(* Logix 5000 project; controller FV vendor 1 type 14 code 217 rev 31.11; software revision 31.00; part 45 of 63 *)
(* tags used below, declared in another part *)
   CWD : CHECKWORD_FLAGS;
   FV_AV1A : PlantItem;   // AV1A
   FV_AV3 : PlantItem;   // AV3
   FV_AV4A : PlantItem;   // AV4A
   FV_B62 : INT[255];   // RESEED FLG
   FV_B72 : INT[255];   // LNCIP FLG
   FV_B72_O_2_OutputBit : BOOL;
   FV_FV10_TTX01_AI : PlantItem;   // FV10_TTX01
   FV_FV11_TTX01_AI : PlantItem;   // FV11_TTX01
   FV_FV12_TTX01_AI : PlantItem;   // FV12_TTX01
   FV_FV13_TTX01_AI : PlantItem;   // FV13_TTX01
   FV_FV14_TTX01_AI : PlantItem;   // FV14_TTX01
   FV_FV15_TTX01_AI : PlantItem;   // FV15_TTX01
   FV_FV16_TTX01_AI : PlantItem;   // FV16_TTX01
   FV_FV17_TTX01_AI : PlantItem;   // FV17_TTX01
   FV_FV18_TTX01_AI : PlantItem;   // FV18_TTX01
   FV_FV19_TTX01_AI : PlantItem;   // FV19_TTX01
   FV_FV1_TTX01_AI : PlantItem;   // FV1_TTX01
   FV_FV20_TTX01_AI : PlantItem;   // FV20_TTX01
   FV_FV21_TTX01_AI : PlantItem;   // FV21_TTX01
   FV_FV22_TTX01_AI : PlantItem;   // FV22_TTX01
   FV_FV23_TTX01_AI : PlantItem;   // FV23_TTX01
   FV_FV24_TTX01_AI : PlantItem;   // FV24_TTX01
   FV_FV25_TTX01_AI : PlantItem;   // FV25_TTX01
   FV_FV26_TTX01_AI : PlantItem;   // FV26_TTX01
   FV_FV26_TTX02_AI : PlantItem;   // FV26_TTX02
   FV_FV27_TTX01_AI : PlantItem;   // FV27_TTX01
   FV_FV27_TTX02_AI : PlantItem;   // FV27_TTX02
   FV_FV28_TTX01_AI : PlantItem;   // FV28_TTX01
   FV_FV28_TTX02_AI : PlantItem;   // FV28_TTX02
   FV_FV29_TTX01_AI : PlantItem;   // FV29_TTX01
   FV_FV29_TTX02_AI : PlantItem;   // FV29_TTX02
   FV_FV2_TTX01_AI : PlantItem;   // FV2_TTX01
   FV_FV30_TTX01_AI : PlantItem;   // FV30_TTX01
   FV_FV30_TTX02_AI : PlantItem;   // FV30_TTX02
   FV_FV31_TTX01_AI : PlantItem;   // FV31_TTX01
   FV_FV31_TTX02_AI : PlantItem;   // FV31_TTX02
   FV_FV3_TTX01_AI : PlantItem;   // FV3_TTX01
   FV_FV4_TTX01_AI : PlantItem;   // FV4_TTX01
   FV_FV5_TTX01_AI : PlantItem;   // FV5_TTX01
   FV_FV6_TTX01_AI : PlantItem;   // FV6_TTX01
   FV_FV7_TTX01_AI : PlantItem;   // FV7_TTX01
   FV_FV8_TTX01_AI : PlantItem;   // FV8_TTX01
   FV_FV9_TTX01_AI : PlantItem;   // FV9_TTX01
   FV_GLYCOL_AI : PlantItem;   // GLYCOL
   FV_N111 : INT[50];   // FV1, CURRENT FV DATA
   FV_N112 : INT[50];   // FV2, CURRENT FV DATA
   FV_N113 : INT[50];   // FV3, CURRENT FV DATA
   FV_N114 : INT[50];   // FV4, CURRENT FV DATA
   FV_N115 : INT[50];   // FV5, CURRENT FV DATA
   FV_N116 : INT[50];   // FV6, CURRENT FV DATA
   FV_N117 : INT[50];   // FV7, CURRENT FV DATA
   FV_N118 : INT[50];   // FV8, CURRENT FV DATA
   FV_N119 : INT[50];   // FV9, CURRENT FV DATA
   FV_N12 : INT[255];   // SYS_PARMS System Parameter Fil e
   FV_N120 : INT[50];   // FV10, CURRENT FV DATA
   FV_N121 : INT[50];   // FV11, CURRENT FV DATA
   FV_N122 : INT[50];   // FV12, CURRENT FV DATA
   FV_N123 : INT[50];   // FV13, CURRENT FV DATA
   FV_N124 : INT[50];   // FV14, CURRENT FV DATA
   FV_N125 : INT[50];   // FV15, CURRENT FV DATA
   FV_N126 : INT[50];   // FV16, CURRENT FV DATA
   FV_N127 : INT[50];   // FV17, CURRENT FV DATA
   FV_N128 : INT[50];   // FV18, CURRENT FV DATA
   FV_N129 : INT[50];   // FV19, CURRENT FV DATA
   FV_N130 : INT[50];   // FV20, CURRENT FV DATA
   FV_N131 : INT[50];   // FV21, CURRENT FV DATA
   FV_N132 : INT[50];   // FV22, CURRENT FV DATA
   FV_N133 : INT[50];   // FV23, CURRENT FV DATA
   FV_N134 : INT[50];   // FV24, CURRENT FV DATA
   FV_N135 : INT[50];   // FV25, CURRENT FV DATA
   FV_N136 : INT[50];   // YSV1, CURRENT FV DATA
   FV_N137 : INT[50];   // YSV2, CURRENT FV DATA
   FV_N138 : INT[50];   // YSV3, CURRENT FV DATA
   FV_N139 : INT[255];   // YST1
   FV_N140 : INT[255];   // YST2
   FV_N141 : INT[255];   // YSV1 DATA
   FV_N142 : INT[255];   // YSV2 DATA
   FV_N143 : INT[255];   // YSV3 DATA
   FV_N146 : INT[50];   // FV26, CURRENT FV DATA
   FV_N147 : INT[50];   // FV27, CURRENT FV DATA
   FV_N148 : INT[50];   // FV28, CURRENT FV DATA
   FV_N149 : INT[50];   // FV29, CURRENT FV DATA
   FV_N150 : INT[50];   // FV30, CURRENT FV DATA
   FV_N151 : INT[50];   // FV31, CURRENT FV DATA
   FV_N7 : INT[255];   // INTEGER
   FV_N70 : INT[255];   // LNCIP <PC
   FV_N71 : INT[255];   // LNCIP >PC
   FV_PX2 : PlantItem;   // PX2
   FV_PX3 : PlantItem;   // PX3
   FV_SOV1 : PlantItem;   // SOV1
   FV_T73 : TIMER[10];
   FV_TTX_YS_001_AI : PlantItem;   // TTX_YS_001
   FV_TTX_YS_002_AI : PlantItem;   // TTX_YS_002
   FV_YSV1_TTX01_AI : PlantItem;   // YSV1_TTX01
   FV_YSV1_WTX01_AI : PlantItem;   // YSV1_WTX01
   FV_YSV2_TTX01_AI : PlantItem;   // YSV2_TTX01
   FV_YSV2_WTX01_AI : PlantItem;   // YSV2_WTX01
   FV_YSV3_TTX01_AI : PlantItem;   // YSV3_TTX01
   FV_YSV3_WTX01_AI : PlantItem;   // YSV3_WTX01
(* FV_Common, continued *)

ROUTINE FV_LNCIP_CP_36   (* ladder *)
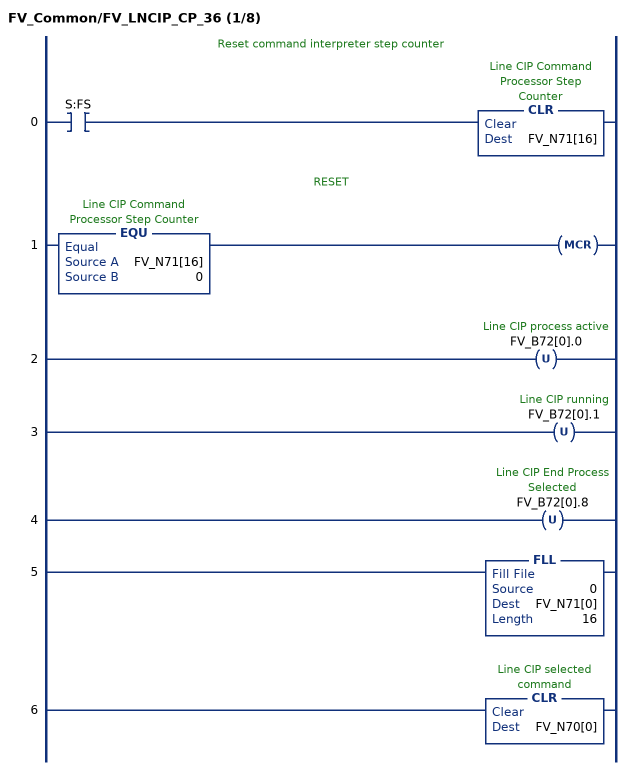
   // Reset command interpreter step counter
   0: XIC(S:FS)CLR(FV_N71[16]);
   // RESET
   1: EQU(FV_N71[16],0)MCR();
   2: OTU(FV_B72[0].0);
   3: OTU(FV_B72[0].1);
   4: OTU(FV_B72[0].8);
   5: FLL(0,FV_N71[0],16);
   6: CLR(FV_N70[0]);
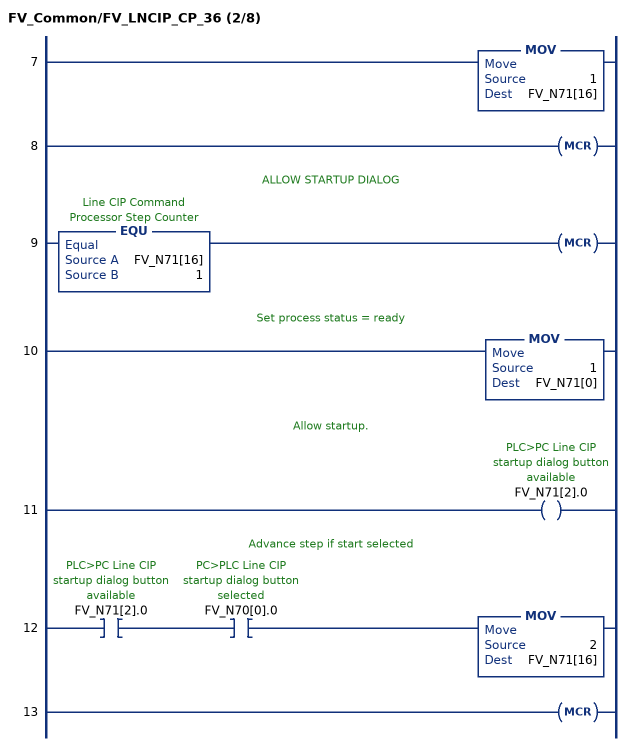
   7: MOV(1,FV_N71[16]);
   8: MCR();
   // ALLOW STARTUP DIALOG
   9: EQU(FV_N71[16],1)MCR();
   // Set process status = ready
   10: MOV(1,FV_N71[0]);
   // Allow startup.
   11: OTE(FV_N71[2].0);
   // Advance step if start selected
   12: XIC(FV_N71[2].0)XIC(FV_N70[0].0)MOV(2,FV_N71[16]);
   13: MCR();
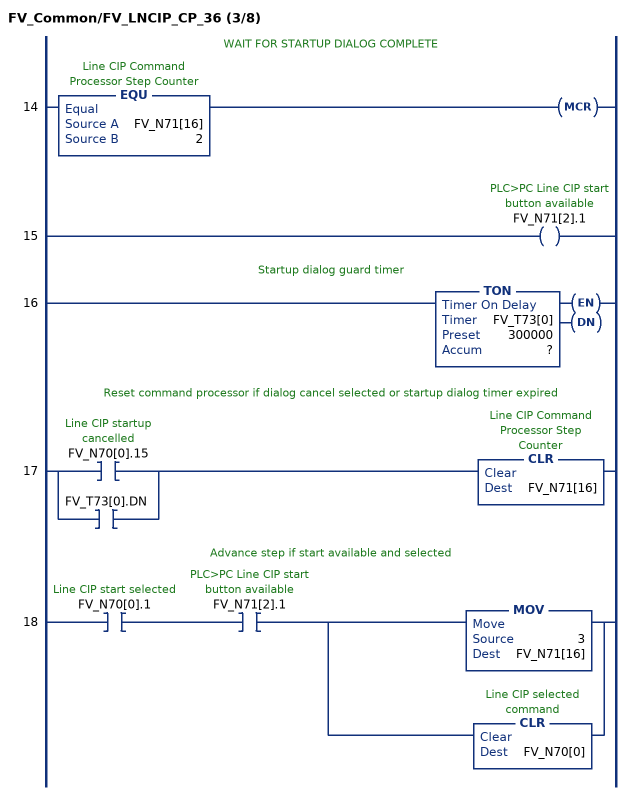
   // WAIT FOR STARTUP DIALOG COMPLETE
   14: EQU(FV_N71[16],2)MCR();
   15: OTE(FV_N71[2].1);
   // Startup dialog guard timer
   16: TON(FV_T73[0],?,?);
   // Reset command processor if dialog cancel selected or startup dialog timer expired
   17: [XIC(FV_N70[0].15) ,XIC(FV_T73[0].DN) ]CLR(FV_N71[16]);
   // Advance step if start available and selected
   18: XIC(FV_N70[0].1)XIC(FV_N71[2].1)[MOV(3,FV_N71[16]) ,CLR(FV_N70[0]) ];
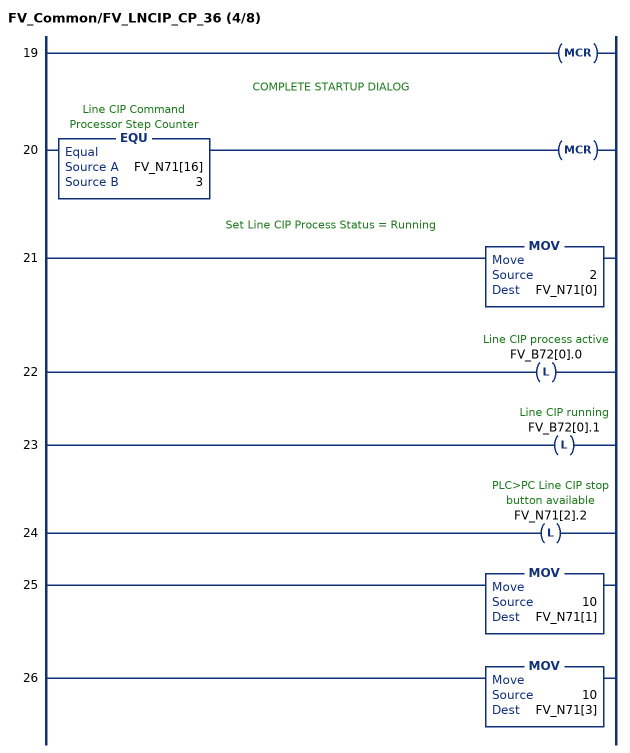
   19: MCR();
   // COMPLETE STARTUP DIALOG
   20: EQU(FV_N71[16],3)MCR();
   // Set Line CIP Process Status = Running
   21: MOV(2,FV_N71[0]);
   22: OTL(FV_B72[0].0);
   23: OTL(FV_B72[0].1);
   24: OTL(FV_N71[2].2);
   25: MOV(10,FV_N71[1]);
   26: MOV(10,FV_N71[3]);
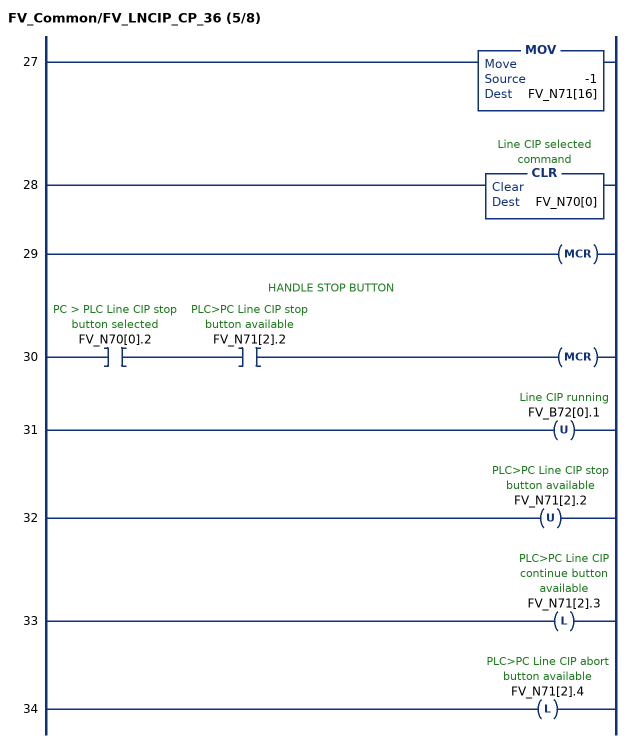
   27: MOV(-1,FV_N71[16]);
   28: CLR(FV_N70[0]);
   29: MCR();
   // HANDLE STOP BUTTON
   30: XIC(FV_N70[0].2)XIC(FV_N71[2].2)MCR();
   31: OTU(FV_B72[0].1);
   32: OTU(FV_N71[2].2);
   33: OTL(FV_N71[2].3);
   34: OTL(FV_N71[2].4);
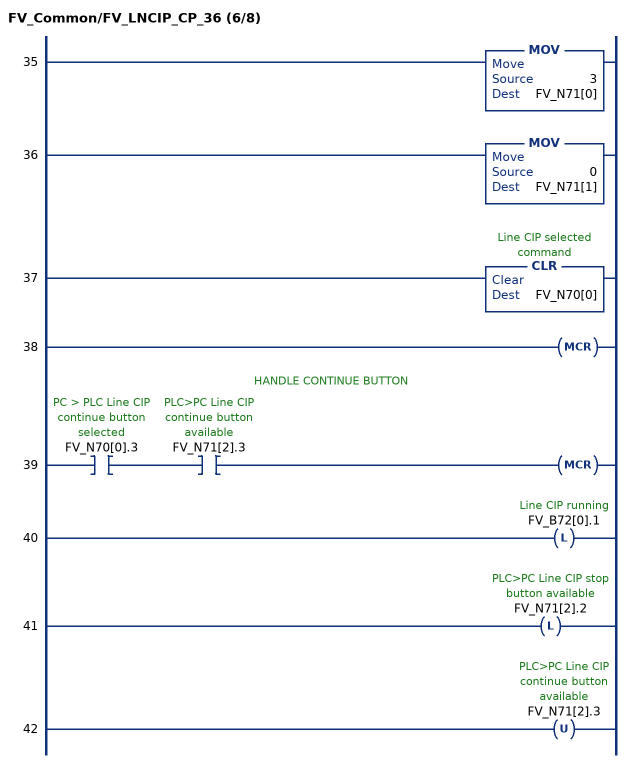
   35: MOV(3,FV_N71[0]);
   36: MOV(0,FV_N71[1]);
   37: CLR(FV_N70[0]);
   38: MCR();
   // HANDLE CONTINUE BUTTON
   39: XIC(FV_N70[0].3)XIC(FV_N71[2].3)MCR();
   40: OTL(FV_B72[0].1);
   41: OTL(FV_N71[2].2);
   42: OTU(FV_N71[2].3);
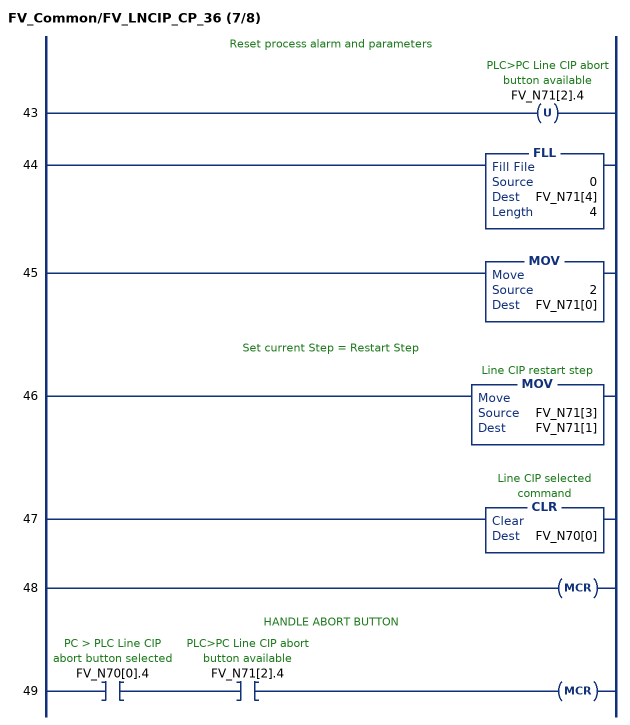
   // Reset process alarm and parameters
   43: OTU(FV_N71[2].4);
   44: FLL(0,FV_N71[4],4);
   45: MOV(2,FV_N71[0]);
   // Set current Step = Restart Step
   46: MOV(FV_N71[3],FV_N71[1]);
   47: CLR(FV_N70[0]);
   48: MCR();
   // HANDLE ABORT BUTTON
   49: XIC(FV_N70[0].4)XIC(FV_N71[2].4)MCR();
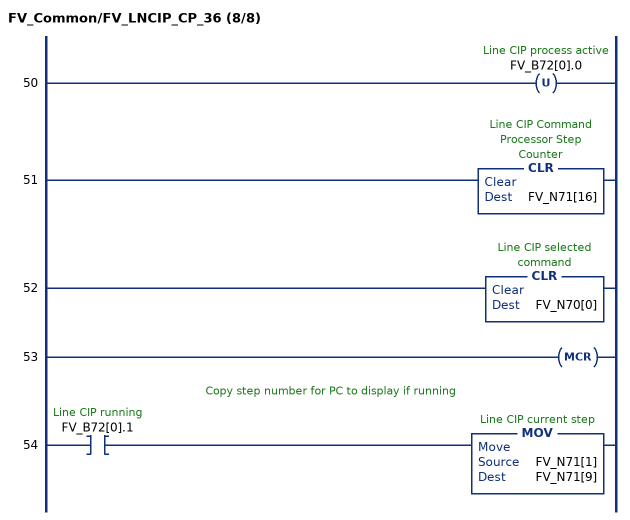
   50: OTU(FV_B72[0].0);
   51: CLR(FV_N71[16]);
   52: CLR(FV_N70[0]);
   53: MCR();
   // Copy step number for PC to display if running
   54: XIC(FV_B72[0].1)MOV(FV_N71[1],FV_N71[9]);
END_ROUTINE

ROUTINE FV_LNCIP_MC_35   (* ladder *)
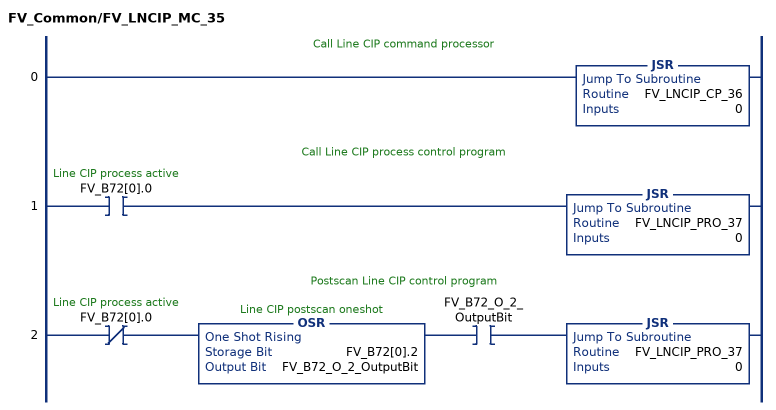
   // Call Line CIP command processor
   0: JSR(FV_LNCIP_CP_36,0);
   // Call Line CIP process control program
   1: XIC(FV_B72[0].0)JSR(FV_LNCIP_PRO_37,0);
   // Postscan Line CIP control program
   2: XIO(FV_B72[0].0)OSR(FV_B72[0].2,FV_B72_O_2_OutputBit)XIC(FV_B72_O_2_OutputBit)JSR(FV_LNCIP_PRO_37,0);
END_ROUTINE

ROUTINE FV_LNCIP_PRO_37   (* ladder *)
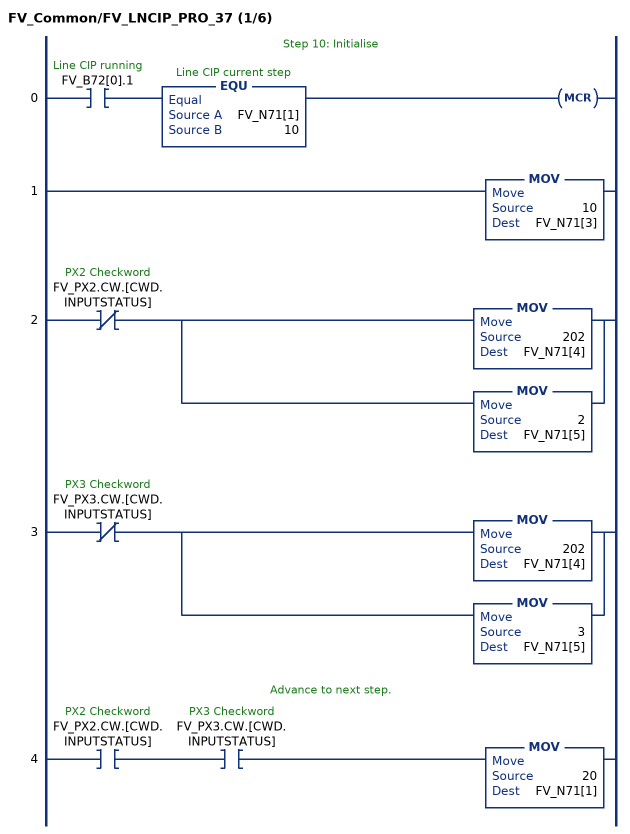
   // Step 10: Initialise
   0: XIC(FV_B72[0].1)EQU(FV_N71[1],10)MCR();
   1: MOV(10,FV_N71[3]);
   2: XIO(FV_PX2.CW.[CWD.INPUTSTATUS])[MOV(202,FV_N71[4]) ,MOV(2,FV_N71[5]) ];
   3: XIO(FV_PX3.CW.[CWD.INPUTSTATUS])[MOV(202,FV_N71[4]) ,MOV(3,FV_N71[5]) ];
   // Advance to next step.
   4: XIC(FV_PX2.CW.[CWD.INPUTSTATUS])XIC(FV_PX3.CW.[CWD.INPUTSTATUS])MOV(20,FV_N71[1]);
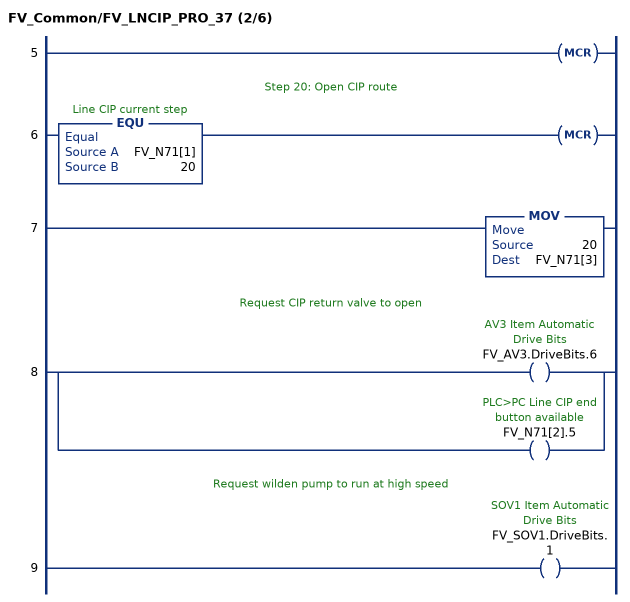
   5: MCR();
   // Step 20: Open CIP route
   6: EQU(FV_N71[1],20)MCR();
   7: MOV(20,FV_N71[3]);
   // Request CIP return valve to open
   8: [OTE(FV_AV3.DriveBits.6) ,OTE(FV_N71[2].5) ];
   // Request wilden pump to run at high speed
   9: OTE(FV_SOV1.DriveBits.1);
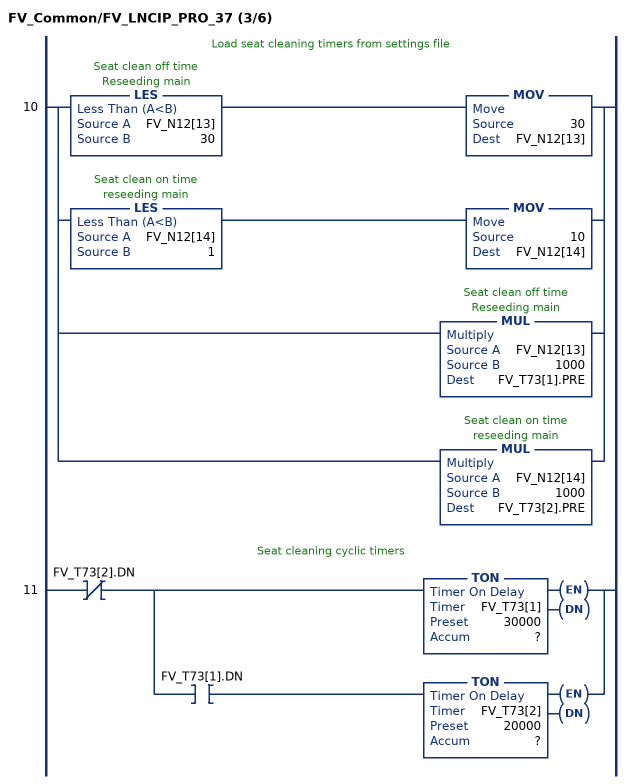
   // Load seat cleaning timers from settings file
   10: [LES(FV_N12[13],30) MOV(30,FV_N12[13]) ,LES(FV_N12[14],1) MOV(10,FV_N12[14]) ,MUL(FV_N12[13],1000,FV_T73[1].PRE) ,MUL(FV_N12[14],1000,FV_T73[2].PRE) ];
   // Seat cleaning cyclic timers
   11: XIO(FV_T73[2].DN)[TON(FV_T73[1],?,?) ,XIC(FV_T73[1].DN) TON(FV_T73[2],?,?) ];
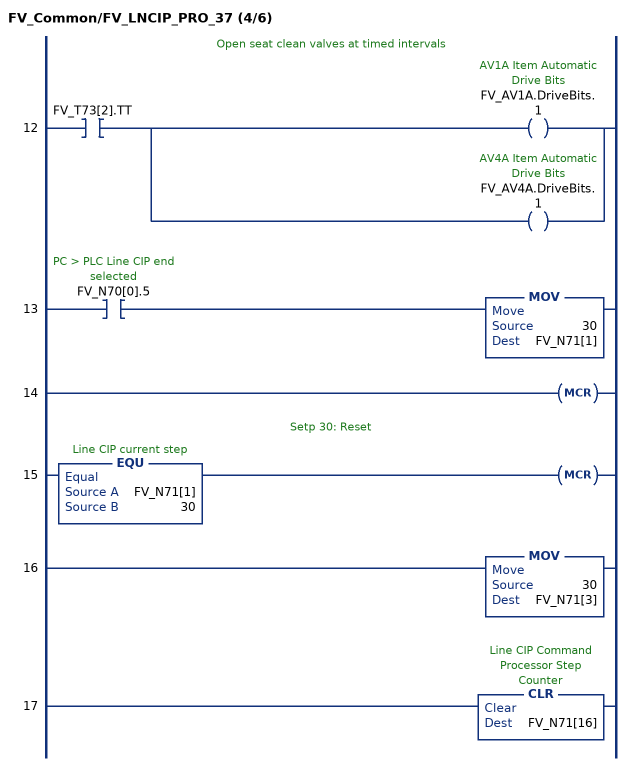
   // Open seat clean valves at timed intervals
   12: XIC(FV_T73[2].TT)[OTE(FV_AV1A.DriveBits.1) ,OTE(FV_AV4A.DriveBits.1) ];
   13: XIC(FV_N70[0].5)MOV(30,FV_N71[1]);
   14: MCR();
   // Setp 30: Reset
   15: EQU(FV_N71[1],30)MCR();
   16: MOV(30,FV_N71[3]);
   17: CLR(FV_N71[16]);
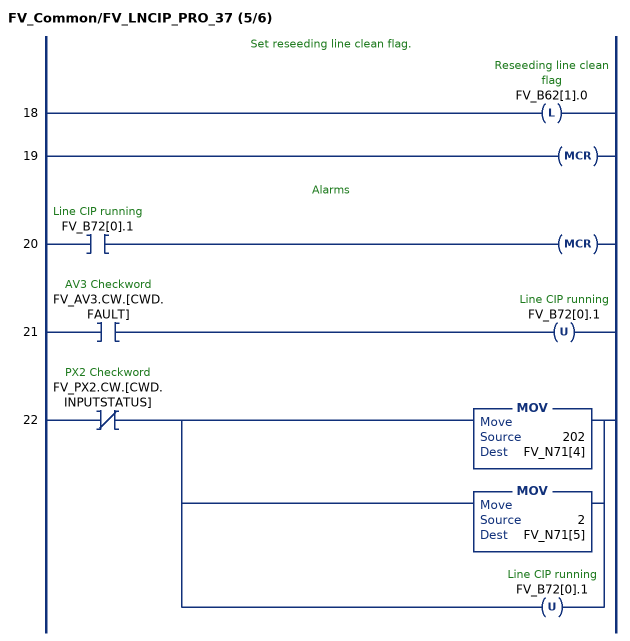
   // Set reseeding line clean flag.
   18: OTL(FV_B62[1].0);
   19: MCR();
   // Alarms
   20: XIC(FV_B72[0].1)MCR();
   21: XIC(FV_AV3.CW.[CWD.FAULT])OTU(FV_B72[0].1);
   22: XIO(FV_PX2.CW.[CWD.INPUTSTATUS])[MOV(202,FV_N71[4]) ,MOV(2,FV_N71[5]) ,OTU(FV_B72[0].1) ];
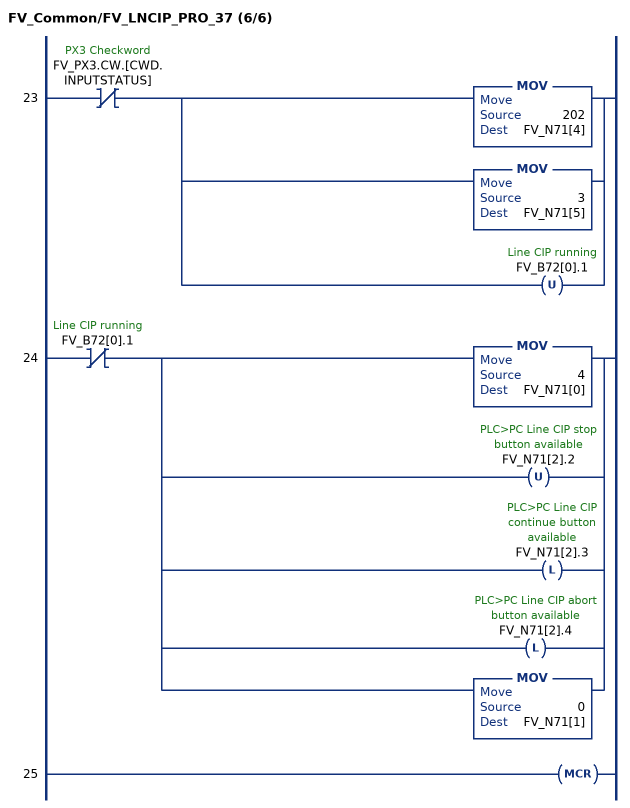
   23: XIO(FV_PX3.CW.[CWD.INPUTSTATUS])[MOV(202,FV_N71[4]) ,MOV(3,FV_N71[5]) ,OTU(FV_B72[0].1) ];
   24: XIO(FV_B72[0].1)[MOV(4,FV_N71[0]) ,OTU(FV_N71[2].2) ,OTL(FV_N71[2].3) ,OTL(FV_N71[2].4) ,MOV(0,FV_N71[1]) ];
   25: MCR();
END_ROUTINE

ROUTINE FV_Move_Temps_To_DataFiles   (* ladder *)
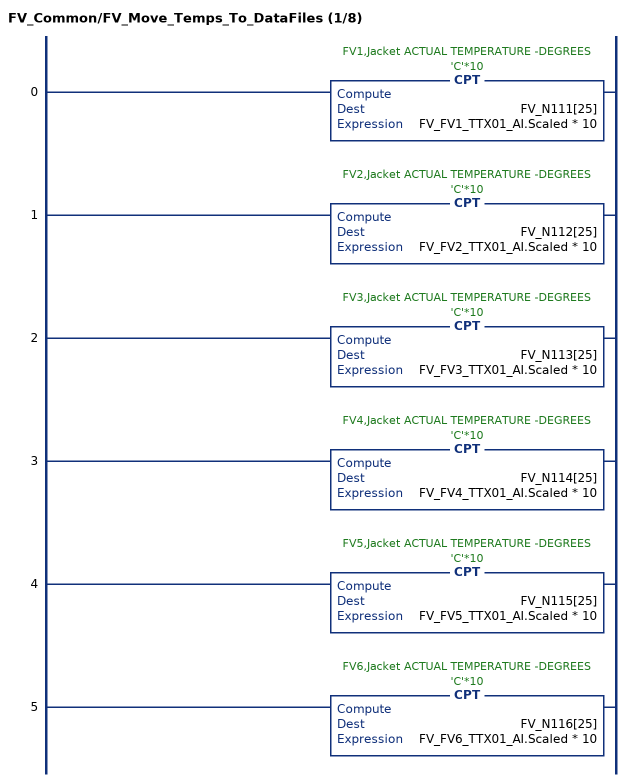
   0: CPT(FV_N111[25],FV_FV1_TTX01_AI.Scaled * 10);
   1: CPT(FV_N112[25],FV_FV2_TTX01_AI.Scaled * 10);
   2: CPT(FV_N113[25],FV_FV3_TTX01_AI.Scaled * 10);
   3: CPT(FV_N114[25],FV_FV4_TTX01_AI.Scaled * 10);
   4: CPT(FV_N115[25],FV_FV5_TTX01_AI.Scaled * 10);
   5: CPT(FV_N116[25],FV_FV6_TTX01_AI.Scaled * 10);
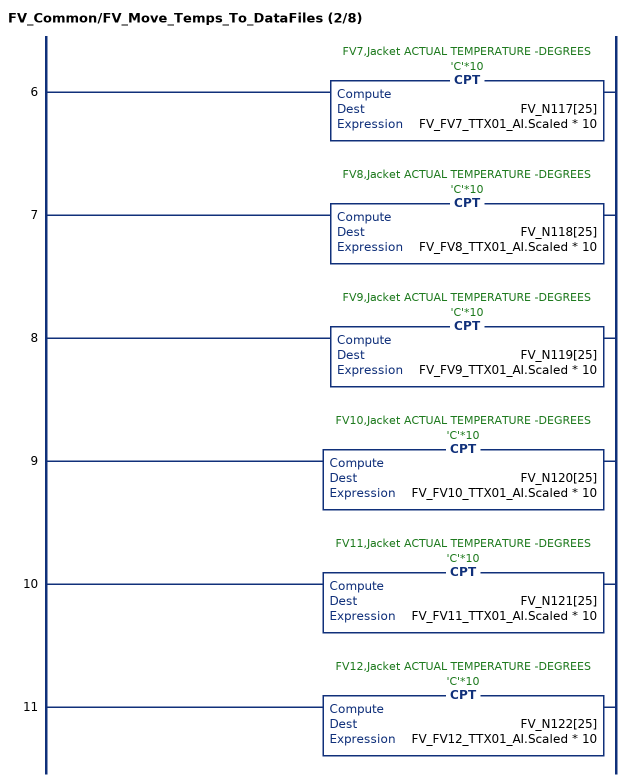
   6: CPT(FV_N117[25],FV_FV7_TTX01_AI.Scaled * 10);
   7: CPT(FV_N118[25],FV_FV8_TTX01_AI.Scaled * 10);
   8: CPT(FV_N119[25],FV_FV9_TTX01_AI.Scaled * 10);
   9: CPT(FV_N120[25],FV_FV10_TTX01_AI.Scaled * 10);
   10: CPT(FV_N121[25],FV_FV11_TTX01_AI.Scaled * 10);
   11: CPT(FV_N122[25],FV_FV12_TTX01_AI.Scaled * 10);
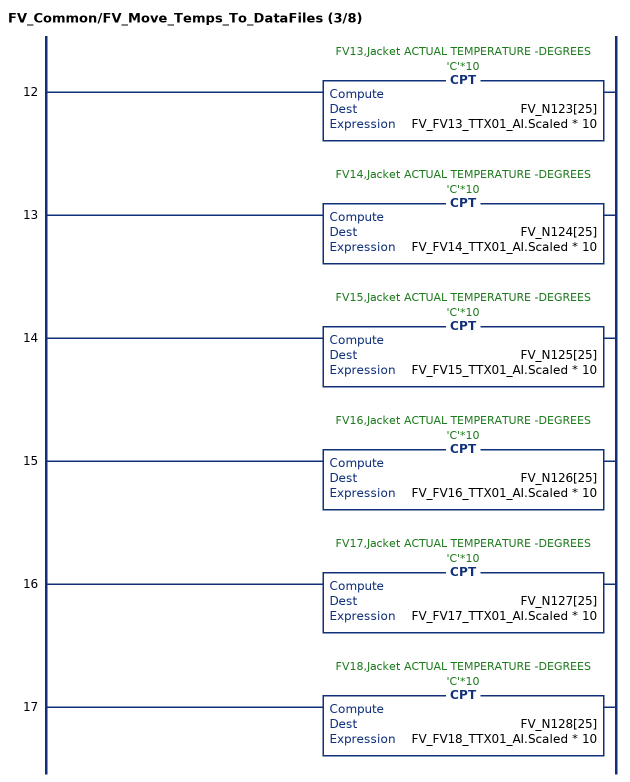
   12: CPT(FV_N123[25],FV_FV13_TTX01_AI.Scaled * 10);
   13: CPT(FV_N124[25],FV_FV14_TTX01_AI.Scaled * 10);
   14: CPT(FV_N125[25],FV_FV15_TTX01_AI.Scaled * 10);
   15: CPT(FV_N126[25],FV_FV16_TTX01_AI.Scaled * 10);
   16: CPT(FV_N127[25],FV_FV17_TTX01_AI.Scaled * 10);
   17: CPT(FV_N128[25],FV_FV18_TTX01_AI.Scaled * 10);
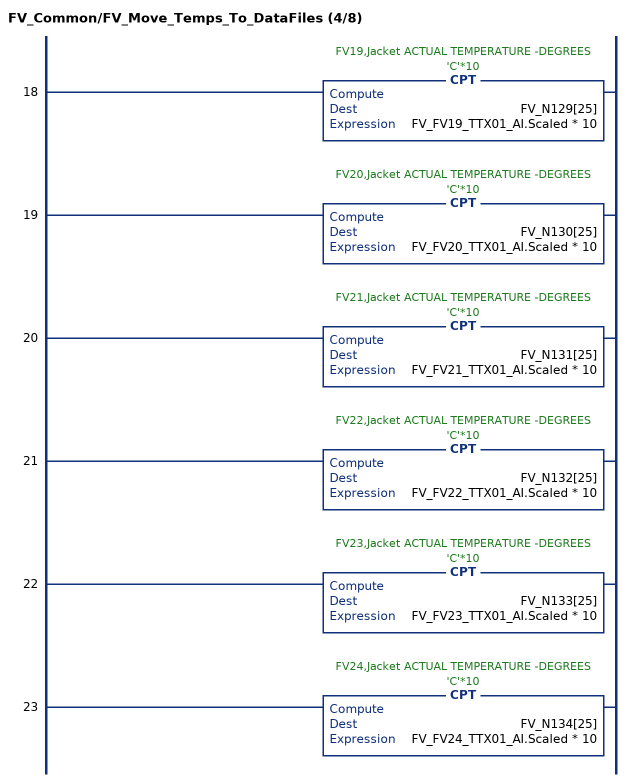
   18: CPT(FV_N129[25],FV_FV19_TTX01_AI.Scaled * 10);
   19: CPT(FV_N130[25],FV_FV20_TTX01_AI.Scaled * 10);
   20: CPT(FV_N131[25],FV_FV21_TTX01_AI.Scaled * 10);
   21: CPT(FV_N132[25],FV_FV22_TTX01_AI.Scaled * 10);
   22: CPT(FV_N133[25],FV_FV23_TTX01_AI.Scaled * 10);
   23: CPT(FV_N134[25],FV_FV24_TTX01_AI.Scaled * 10);
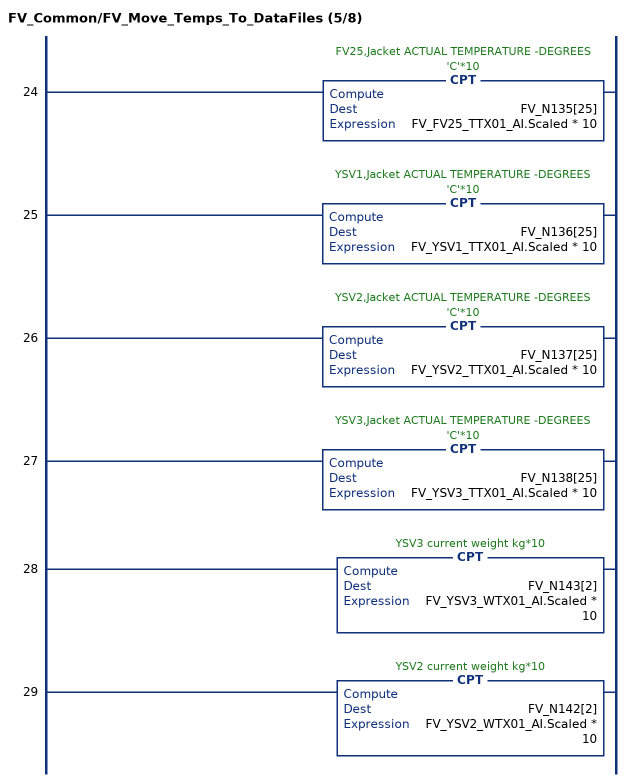
   24: CPT(FV_N135[25],FV_FV25_TTX01_AI.Scaled * 10);
   25: CPT(FV_N136[25],FV_YSV1_TTX01_AI.Scaled * 10);
   26: CPT(FV_N137[25],FV_YSV2_TTX01_AI.Scaled * 10);
   27: CPT(FV_N138[25],FV_YSV3_TTX01_AI.Scaled * 10);
   28: CPT(FV_N143[2],FV_YSV3_WTX01_AI.Scaled * 10);
   29: CPT(FV_N142[2],FV_YSV2_WTX01_AI.Scaled * 10);
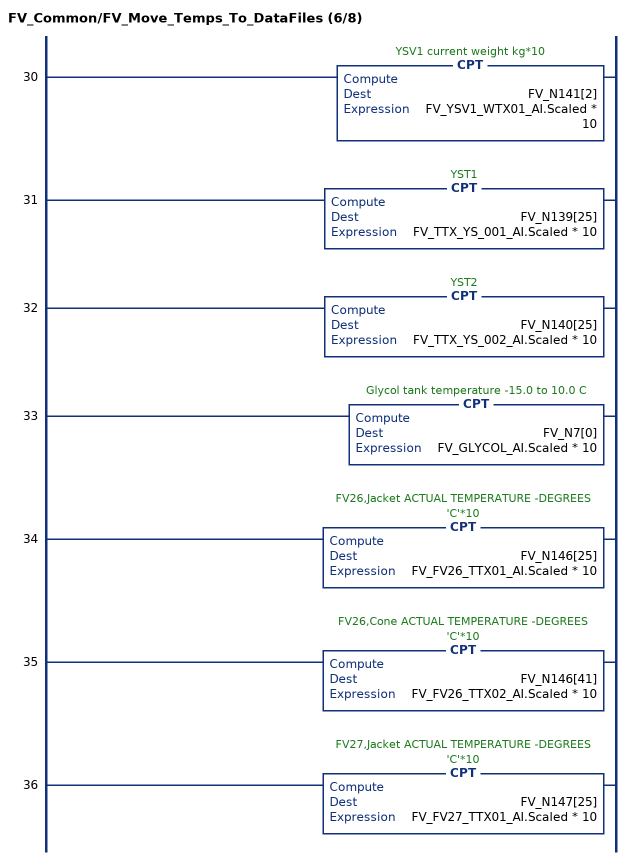
   30: CPT(FV_N141[2],FV_YSV1_WTX01_AI.Scaled * 10);
   31: CPT(FV_N139[25],FV_TTX_YS_001_AI.Scaled * 10);
   32: CPT(FV_N140[25],FV_TTX_YS_002_AI.Scaled * 10);
   33: CPT(FV_N7[0],FV_GLYCOL_AI.Scaled * 10);
   34: CPT(FV_N146[25],FV_FV26_TTX01_AI.Scaled * 10);
   35: CPT(FV_N146[41],FV_FV26_TTX02_AI.Scaled * 10);
   36: CPT(FV_N147[25],FV_FV27_TTX01_AI.Scaled * 10);
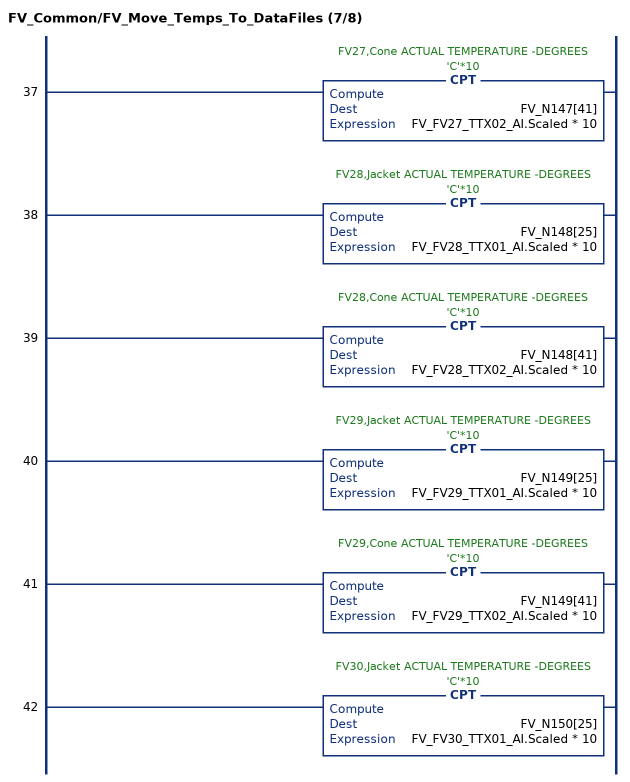
   37: CPT(FV_N147[41],FV_FV27_TTX02_AI.Scaled * 10);
   38: CPT(FV_N148[25],FV_FV28_TTX01_AI.Scaled * 10);
   39: CPT(FV_N148[41],FV_FV28_TTX02_AI.Scaled * 10);
   40: CPT(FV_N149[25],FV_FV29_TTX01_AI.Scaled * 10);
   41: CPT(FV_N149[41],FV_FV29_TTX02_AI.Scaled * 10);
   42: CPT(FV_N150[25],FV_FV30_TTX01_AI.Scaled * 10);
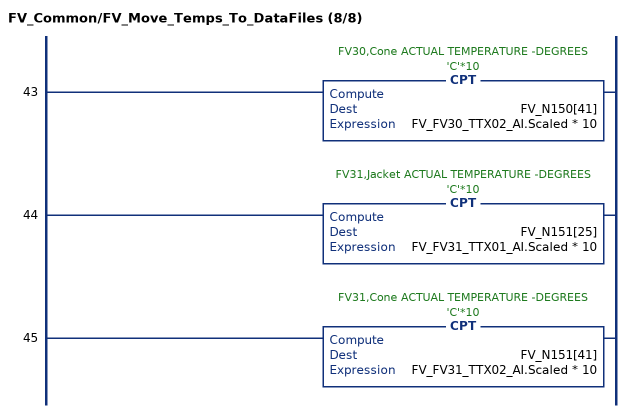
   43: CPT(FV_N150[41],FV_FV30_TTX02_AI.Scaled * 10);
   44: CPT(FV_N151[25],FV_FV31_TTX01_AI.Scaled * 10);
   45: CPT(FV_N151[41],FV_FV31_TTX02_AI.Scaled * 10);
END_ROUTINE
